REGION Network 5: Transfering
   RUNG wire#powerrail
      Contact( "R-201_Write_TO_T-102_DB".Transfering )
      Coil( "T-102_Read_FROM_R-201_DB".Transfering )
   END_RUNG
   // the same network as SCL:
   "T-102_Read_FROM_R-201_DB".Transfering := "R-201_Write_TO_T-102_DB".Transfering;
END_REGION

REGION Network 6: Filling Done
   RUNG wire#powerrail
      Contact( "R-201_Write_TO_T-102_DB".FillingDone )
      Coil( "T-102_Read_FROM_R-201_DB".FillingDone )
   END_RUNG
   // the same network as SCL:
   "T-102_Read_FROM_R-201_DB".FillingDone := "R-201_Write_TO_T-102_DB".FillingDone;
END_REGION

REGION Network 7: Aborting
   RUNG wire#powerrail
      Contact( "R-201_Write_TO_T-102_DB".Abort )
      Coil( "T-102_Read_FROM_R-201_DB".Aborting )
   END_RUNG
   // the same network as SCL:
   "T-102_Read_FROM_R-201_DB".Aborting := "R-201_Write_TO_T-102_DB".Abort;
END_REGION

REGION Network 8: Release Tank
   RUNG wire#powerrail
      Contact( "R-201_Write_TO_T-102_DB".ReleaseTank )
      Coil( "T-102_Read_FROM_R-201_DB".ReleaseTank )
   END_RUNG
   // the same network as SCL:
   "T-102_Read_FROM_R-201_DB".ReleaseTank := "R-201_Write_TO_T-102_DB".ReleaseTank;
END_REGION
END_FUNCTION

// folder: State MACHINE/1)Tanks/Tank T-102 (Y)/T-102 <---> R-202

FUNCTION "T-102_Signals_FROM_R-202" : Void   // FC70, LAD
{ S7_Optimized_Access := 'TRUE' }
VERSION : 0.1
BEGIN

REGION Network 1: Start Pouring Sequence
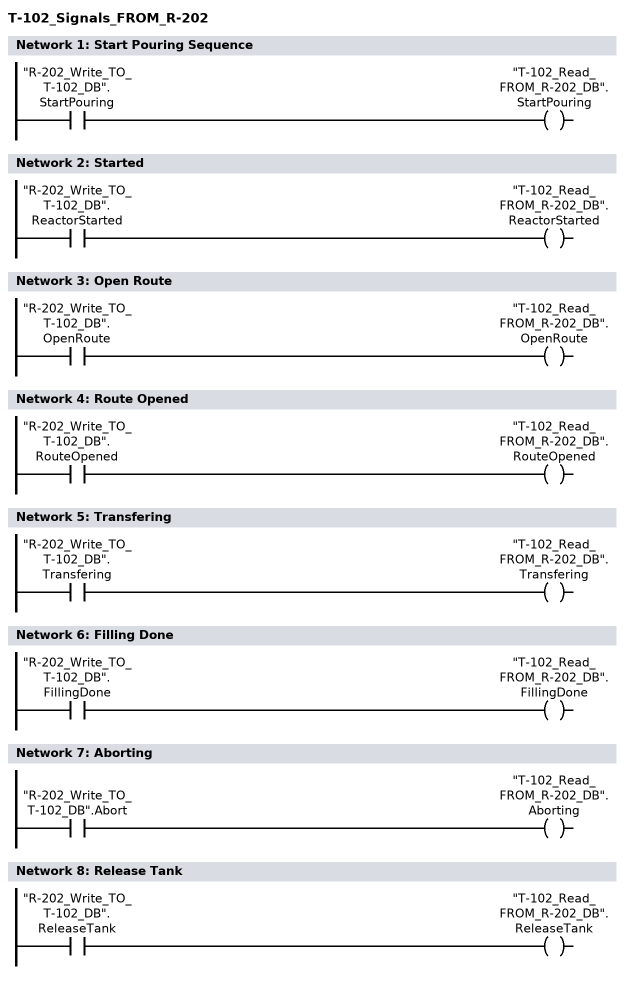
   RUNG wire#powerrail
      Contact( "R-202_Write_TO_T-102_DB".StartPouring )
      Coil( "T-102_Read_FROM_R-202_DB".StartPouring )
   END_RUNG
   // the same network as SCL:
   "T-102_Read_FROM_R-202_DB".StartPouring := "R-202_Write_TO_T-102_DB".StartPouring;
END_REGION

REGION Network 2: Started
   RUNG wire#powerrail
      Contact( "R-202_Write_TO_T-102_DB".ReactorStarted )
      Coil( "T-102_Read_FROM_R-202_DB".ReactorStarted )
   END_RUNG
   // the same network as SCL:
   "T-102_Read_FROM_R-202_DB".ReactorStarted := "R-202_Write_TO_T-102_DB".ReactorStarted;
END_REGION

REGION Network 3: Open Route
   RUNG wire#powerrail
      Contact( "R-202_Write_TO_T-102_DB".OpenRoute )
      Coil( "T-102_Read_FROM_R-202_DB".OpenRoute )
   END_RUNG
   // the same network as SCL:
   "T-102_Read_FROM_R-202_DB".OpenRoute := "R-202_Write_TO_T-102_DB".OpenRoute;
END_REGION

REGION Network 4: Route Opened
   RUNG wire#powerrail
      Contact( "R-202_Write_TO_T-102_DB".RouteOpened )
      Coil( "T-102_Read_FROM_R-202_DB".RouteOpened )
   END_RUNG
   // the same network as SCL:
   "T-102_Read_FROM_R-202_DB".RouteOpened := "R-202_Write_TO_T-102_DB".RouteOpened;
END_REGION

REGION Network 5: Transfering
   RUNG wire#powerrail
      Contact( "R-202_Write_TO_T-102_DB".Transfering )
      Coil( "T-102_Read_FROM_R-202_DB".Transfering )
   END_RUNG
   // the same network as SCL:
   "T-102_Read_FROM_R-202_DB".Transfering := "R-202_Write_TO_T-102_DB".Transfering;
END_REGION

REGION Network 6: Filling Done
   RUNG wire#powerrail
      Contact( "R-202_Write_TO_T-102_DB".FillingDone )
      Coil( "T-102_Read_FROM_R-202_DB".FillingDone )
   END_RUNG
   // the same network as SCL:
   "T-102_Read_FROM_R-202_DB".FillingDone := "R-202_Write_TO_T-102_DB".FillingDone;
END_REGION

REGION Network 7: Aborting
   RUNG wire#powerrail
      Contact( "R-202_Write_TO_T-102_DB".Abort )
      Coil( "T-102_Read_FROM_R-202_DB".Aborting )
   END_RUNG
   // the same network as SCL:
   "T-102_Read_FROM_R-202_DB".Aborting := "R-202_Write_TO_T-102_DB".Abort;
END_REGION

REGION Network 8: Release Tank
   RUNG wire#powerrail
      Contact( "R-202_Write_TO_T-102_DB".ReleaseTank )
      Coil( "T-102_Read_FROM_R-202_DB".ReleaseTank )
   END_RUNG
   // the same network as SCL:
   "T-102_Read_FROM_R-202_DB".ReleaseTank := "R-202_Write_TO_T-102_DB".ReleaseTank;
END_REGION
END_FUNCTION

// folder: State MACHINE/1)Tanks/Tank T-102 (Y)/T-102 <---> T-104

FUNCTION "T-102_Signals_FROM_T-104" : Void   // FC55, LAD
{ S7_Optimized_Access := 'TRUE' }
VERSION : 0.1
BEGIN

REGION Network 1: Start Sequence
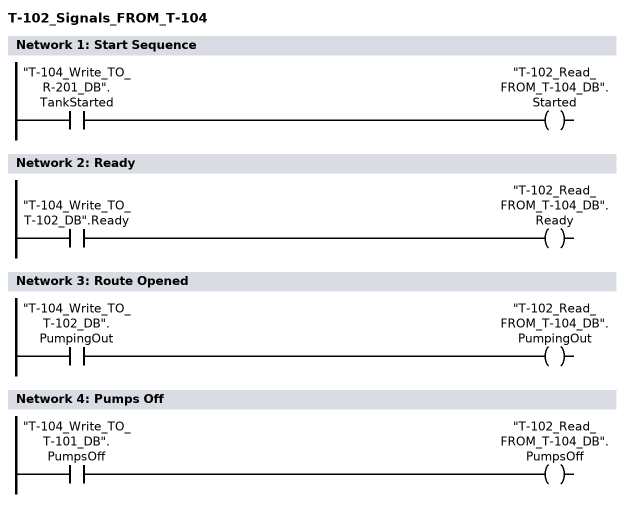
   RUNG wire#powerrail
      Contact( "T-104_Write_TO_R-201_DB".TankStarted )
      Coil( "T-102_Read_FROM_T-104_DB".Started )
   END_RUNG
   // the same network as SCL:
   "T-102_Read_FROM_T-104_DB".Started := "T-104_Write_TO_R-201_DB".TankStarted;
END_REGION

REGION Network 2: Ready
   RUNG wire#powerrail
      Contact( "T-104_Write_TO_T-102_DB".Ready )
      Coil( "T-102_Read_FROM_T-104_DB".Ready )
   END_RUNG
   // the same network as SCL:
   "T-102_Read_FROM_T-104_DB".Ready := "T-104_Write_TO_T-102_DB".Ready;
END_REGION

REGION Network 3: Route Opened
   RUNG wire#powerrail
      Contact( "T-104_Write_TO_T-102_DB".PumpingOut )
      Coil( "T-102_Read_FROM_T-104_DB".PumpingOut )
   END_RUNG
   // the same network as SCL:
   "T-102_Read_FROM_T-104_DB".PumpingOut := "T-104_Write_TO_T-102_DB".PumpingOut;
END_REGION

REGION Network 4: Pumps Off
   RUNG wire#powerrail
      Contact( "T-104_Write_TO_T-101_DB".PumpsOff )
      Coil( "T-102_Read_FROM_T-104_DB".PumpsOff )
   END_RUNG
   // the same network as SCL:
   "T-102_Read_FROM_T-104_DB".PumpsOff := "T-104_Write_TO_T-101_DB".PumpsOff;
END_REGION
END_FUNCTION

// folder: State MACHINE/1)Tanks/Tank T-103 (Cooling Tank)

FUNCTION_BLOCK "T-103_SEQ"   // FB33, GRAPH_PLUS
{ S7_Optimized_Access := 'TRUE' }
VERSION : 0.1
   VAR_INPUT
      OFF_SQ : Bool := false;   // Turn sequence off
      INIT_SQ : Bool := false;   // Set sequence to initial state
      ACK_EF : Bool := false;   // Acknowledge all errors and faults
   END_VAR
   VAR_OUTPUT
      S_NO : Int := 0;   // Step number
      S_MORE : Bool := false;   // More steps are available and can be shown in S_NO
      S_ACTIVE : Bool := false;   // Step indicated in S_NO is active
      ERR_FLT : Bool := false;   // Interlock or supervision group error
      AUTO_ON : Bool := false;   // Automatic mode is active
   END_VAR
   VAR
      STATE : Int;   // Current Step in Sequence
      Tank : Struct   // Reactor Ctrl
         IDLE : Bool;
         INITIALIZATION : Bool;   // Sequence initialization
         START : Bool;
         DONE_REACTING : Bool;
         COMPLETE : Bool;   // Reactor Complete Read only
         PARA : Bool;   // PARA load Batch side button
         ABORTING : Bool;   // Sequence about
         WAIT : Bool;   // Wating for Permissive read only
      END_STRUCT;
      TEMP : Struct
         TANKS_BATCH : Real;
         "EMPTY_LV_0%" : Real;
         "MIN_LV_20%" : Real;
         "MAX_LV_80%" : Real;
         "BELOW_32%" : Real;
         "Greater_8%" : Real;
         "PRE-ADD" : Real;
         X_SOL_SIZE : Real;
         Y_SOL_SIZE : Real;
         OFFSEt : Struct
            MAX : Real;
            MIN : Real;
         END_STRUCT;
      END_STRUCT;
      HMI_INFO : Array[0..12] of UInt;
      IF_PAR : G7_IfParPlus_V6;
      RT_DATA : G7_RTDataPlus_V6;   // Internal data area
      Abort : G7_TransitionPlus_V6;   // Transition structure
      Initialize : G7_TransitionPlus_V6;   // Transition structure
      Block : G7_TransitionPlus_V6;   // Transition structure
      Rdy : G7_TransitionPlus_V6;   // Transition structure
      Receive : G7_TransitionPlus_V6;   // Transition structure
      Centrifuge : G7_TransitionPlus_V6;   // Transition structure
      OpenR : G7_TransitionPlus_V6;   // Transition structure
      MinLevel : G7_TransitionPlus_V6;   // Transition structure
      DnTransf : G7_TransitionPlus_V6;   // Transition structure
      Cold : G7_TransitionPlus_V6;   // Transition structure
      POff : G7_TransitionPlus_V6;   // Transition structure
      ClsR : G7_TransitionPlus_V6;   // Transition structure
      DnClng : G7_TransitionPlus_V6;   // Transition structure
      TrSt : G7_TransitionPlus_V6;   // Transition structure
      ROpn : G7_TransitionPlus_V6;   // Transition structure
      Tng : G7_TransitionPlus_V6;   // Transition structure
      ClsFR : G7_TransitionPlus_V6;   // Transition structure
      DnT : G7_TransitionPlus_V6;   // Transition structure
      Init : G7_TransitionPlus_V6;   // Transition structure
      SAut : G7_TransitionPlus_V6;   // Transition structure
      SIn : G7_TransitionPlus_V6;   // Transition structure
      Initd : G7_TransitionPlus_V6;   // Transition structure
      BskFull : G7_TransitionPlus_V6;   // Transition structure
      FeelerRet : G7_TransitionPlus_V6;   // Transition structure
      Ab : G7_TransitionPlus_V6;   // Transition structure
      AbortOn : G7_TransitionPlus_V6;   // Transition structure
      DneAbort : G7_TransitionPlus_V6;   // Transition structure
      Idle : G7_StepPlus_V6;   // Step structure
      Ready : G7_StepPlus_V6;   // Step structure
      SelectSeq : G7_StepPlus_V6;   // Step structure
      Started : G7_StepPlus_V6;   // Step structure
      Filling : G7_StepPlus_V6;   // Step structure
      "Filling/Tansfer" : G7_StepPlus_V6;   // Step structure
      Wait_Temp : G7_StepPlus_V6;   // Step structure
      PmpOff : G7_StepPlus_V6;   // Step structure
      CloseRecirc : G7_StepPlus_V6;   // Step structure
      "USER Ready" : G7_StepPlus_V6;   // Step structure
      ReadyToTransf : G7_StepPlus_V6;   // Step structure
      RouteOpened : G7_StepPlus_V6;   // Step structure
      Transfering : G7_StepPlus_V6;   // Step structure
      CloseFeedRoute : G7_StepPlus_V6;   // Step structure
      DoneTrnf : G7_StepPlus_V6;   // Step structure
      Idle_Init : G7_StepPlus_V6;   // Step structure
      SetAuto : G7_StepPlus_V6;   // Step structure
      SetInitial : G7_StepPlus_V6;   // Step structure
      Done_Init : G7_StepPlus_V6;   // Step structure
      AbortStarting : G7_StepPlus_V6;   // Step structure
      Aborting : G7_StepPlus_V6;   // Step structure
      Abort_Done : G7_StepPlus_V6;   // Step structure
      SINI : Array[0..5] of USInt;
      LSTT : Array[0..26] of USInt;
      ATAJ : Array[0..26] of USInt;
      ATAB : Array[0..26] of USInt;
      PSTT : Array[0..26] of USInt;
      NSTT : Array[0..26] of USInt;
      ASSJ : Array[0..21] of USInt;
      ASSB : Array[0..21] of USInt;
      PTTS : Array[0..21] of USInt;
      NTTS : Array[0..21] of USInt;
      SW_SQTS : Array[0..21] of USInt;
      SWITCH : Array[0..6] of USInt;
      TVX : Array[0..13] of USInt;
      TTX : Array[0..13] of USInt;
      TSX : Array[0..5] of USInt;
      S00X : Array[0..5] of USInt;
      SOFFX : Array[0..5] of USInt;
      SONX : Array[0..5] of USInt;
      SAX : Array[0..5] of USInt;
      SERRX : Array[0..22] of USInt;
      SMX : Array[0..22] of USInt;
      S0X : Array[0..22] of USInt;
      S1X : Array[0..22] of USInt;
      IL_ALARM_INST : Diag_Alarm;
      SUP_ALARM_INST : Diag_Alarm;
      STEP_TIME_ALARM_INST : Diag_Alarm;
      IEC_TIMER_INST : IEC_TIMER;
      TRANSACTION_FLAG : Bool := false;
   END_VAR
   VAR CONSTANT
      "Single R-201 T-101 seq done" : Int := 214;
      "Single R-201 T-102 seq done" : Int := 218;
   END_VAR
   // SINI[0] := 2;
   // LSTT[0] := 19;
   // NSTT[0] := 19;
   // PTTS[0] := 255;
   // TVX[0] := 16#1;
   // TTX[0] := 16#1;
   // TSX[0] := 16#1;
   // S00X[0] := 16#1;
   // SOFFX[0] := 16#1;
   // SONX[0] := 16#1;
   // SAX[0] := 16#1;
   // SERRX[0] := 16#1;
   // SMX[0] := 16#1;
   // S0X[0] := 16#1;
   // S1X[0] := 16#1;
   // LSTT[1] := 15;
   // LSTT[2] := 255;
   // LSTT[3] := 255;
   // LSTT[4] := 3;
   // LSTT[5] := 10;
   // LSTT[6] := 255;
   // LSTT[7] := 255;
   // LSTT[8] := 255;
   // LSTT[9] := 255;
   // LSTT[10] := 255;
   // LSTT[11] := 255;
   // LSTT[21] := 1;
   // LSTT[13] := 255;
   // LSTT[14] := 255;
   // LSTT[15] := 255;
   // LSTT[16] := 255;
   // LSTT[20] := 255;
   // LSTT[23] := 10;
   // LSTT[19] := 255;
   // LSTT[22] := 10;
   // ATAJ[1] := 1;
   // ATAJ[2] := 2;
   // ATAJ[3] := 3;
   // ATAJ[4] := 4;
   // ATAJ[5] := 5;
   // ATAJ[6] := 6;
   // ATAJ[7] := 7;
   // ATAJ[8] := 8;
   // ATAJ[9] := 9;
   // ATAJ[10] := 10;
   // ATAJ[11] := 11;
   // ATAJ[12] := 12;
   // ATAJ[13] := 13;
   // ATAJ[14] := 14;
   // ATAJ[15] := 15;
   // ATAJ[16] := 16;
   // ATAJ[17] := 17;
   // ATAJ[18] := 18;
   // ATAJ[19] := 19;
   // ATAJ[20] := 20;
   // ATAJ[21] := 21;
   // ATAJ[22] := 22;
   // ATAJ[23] := 23;
   // ATAJ[24] := 24;
   // ATAB[1] := 2;
   // ATAB[10] := 10;
   // ATAB[3] := 3;
   // ATAB[4] := 5;
   // ATAB[5] := 4;
   // ATAB[6] := 6;
   // ATAB[7] := 7;
   // ATAB[8] := 8;
   // ATAB[12] := 12;
   // ATAB[11] := 11;
   // ATAB[13] := 13;
   // ATAB[14] := 14;
   // ATAB[15] := 22;
   // ATAB[16] := 16;
   // ATAB[17] := 17;
   // ATAB[18] := 18;
   // ATAB[21] := 21;
   // ATAB[22] := 23;
   // ATAB[23] := 15;
   // ATAB[24] := 24;
   // ATAB[0] := 1;
   // PSTT[10] := 7;
   // PSTT[16] := 13;
   // PSTT[3] := 1;
   // PSTT[4] := 2;
   // PSTT[5] := 2;
   // PSTT[6] := 3;
   // PSTT[7] := 4;
   // PSTT[12] := 9;
   // PSTT[11] := 8;
   // PSTT[13] := 10;
   // PSTT[14] := 11;
   // PSTT[17] := 14;
   // PSTT[18] := 15;
   // PSTT[19] := 16;
   // PSTT[20] := 17;
   // PSTT[21] := 18;
   // PSTT[22] := 12;
   // PSTT[23] := 12;
   // PSTT[24] := 19;
   // NSTT[1] := 15;
   // NSTT[2] := 1;
   // NSTT[3] := 2;
   // NSTT[4] := 3;
   // NSTT[5] := 10;
   // NSTT[6] := 4;
   // NSTT[7] := 5;
   // NSTT[8] := 6;
   // NSTT[9] := 7;
   // NSTT[10] := 8;
   // NSTT[11] := 9;
   // NSTT[21] := 1;
   // NSTT[13] := 11;
   // NSTT[14] := 12;
   // NSTT[15] := 13;
   // NSTT[16] := 14;
   // NSTT[20] := 18;
   // NSTT[23] := 10;
   // NSTT[19] := 17;
   // NSTT[22] := 10;
   // ASSJ[1] := 1;
   // ASSJ[2] := 2;
   // ASSJ[3] := 3;
   // ASSJ[4] := 4;
   // ASSJ[5] := 5;
   // ASSJ[6] := 6;
   // ASSJ[7] := 7;
   // ASSJ[8] := 8;
   // ASSJ[9] := 9;
   // ASSJ[10] := 10;
   // ASSJ[11] := 11;
   // ASSJ[12] := 12;
   // ASSJ[13] := 13;
   // ASSJ[14] := 14;
   // ASSJ[15] := 15;
   // ASSJ[16] := 16;
   // ASSJ[17] := 17;
   // ASSJ[18] := 18;
   // ASSJ[19] := 19;
   // ASSJ[20] := 20;
   // ASSJ[21] := 21;
   // ASSB[1] := 1;
   // ASSB[2] := 2;
   // ASSB[3] := 3;
   // ASSB[4] := 4;
   // ASSB[5] := 5;
   // ASSB[6] := 6;
   // ASSB[7] := 7;
   // ASSB[8] := 8;
   // ASSB[9] := 9;
   // ASSB[10] := 10;
   // ASSB[11] := 11;
   // ASSB[12] := 12;
   // ASSB[13] := 13;
   // ASSB[14] := 14;
   // ASSB[15] := 15;
   // ASSB[16] := 16;
   // ASSB[17] := 17;
   // ASSB[18] := 18;
   // ASSB[19] := 19;
   // ASSB[20] := 20;
   // ASSB[21] := 21;
   // PTTS[4] := 6;
   // PTTS[3] := 255;
   // PTTS[5] := 7;
   // PTTS[6] := 8;
   // PTTS[7] := 9;
   // PTTS[8] := 10;
   // PTTS[9] := 11;
   // PTTS[10] := 255;
   // PTTS[11] := 13;
   // PTTS[12] := 14;
   // PTTS[13] := 15;
   // PTTS[14] := 16;
   // PTTS[15] := 255;
   // PTTS[16] := 18;
   // PTTS[17] := 19;
   // PTTS[18] := 20;
   // PTTS[19] := 255;
   // PTTS[20] := 24;
   // PTTS[21] := 25;
   // SW_SQTS[4] := 2;
   // NTTS[2] := 4;
   // NTTS[3] := 6;
   // NTTS[4] := 7;
   // NTTS[5] := 8;
   // NTTS[6] := 9;
   // NTTS[7] := 10;
   // NTTS[8] := 11;
   // NTTS[9] := 12;
   // NTTS[10] := 13;
   // NTTS[11] := 14;
   // NTTS[12] := 15;
   // NTTS[13] := 16;
   // NTTS[14] := 17;
   // NTTS[15] := 18;
   // NTTS[16] := 19;
   // NTTS[17] := 20;
   // NTTS[18] := 21;
   // NTTS[19] := 24;
   // NTTS[20] := 25;
   // NTTS[21] := 26;
   // SW_SQTS[5] := 2;
   // SW_SQTS[8] := 2;
   // SW_SQTS[9] := 2;
   // SW_SQTS[10] := 3;
   // SW_SQTS[11] := 3;
   // SW_SQTS[12] := 3;
   // SW_SQTS[13] := 4;
   // SW_SQTS[14] := 4;
   // SW_SQTS[15] := 5;
   // SW_SQTS[16] := 5;
   // SW_SQTS[17] := 5;
   // SW_SQTS[18] := 5;
   // SW_SQTS[19] := 6;
   // SW_SQTS[20] := 6;
   // SW_SQTS[21] := 6;
   // SWITCH[3] := 124;
   // SWITCH[0] := 124;
   // SWITCH[2] := 254;
   // SWITCH[4] := 254;
   // PTTS[2] := 3;
   // SW_SQTS[3] := 2;
   // SWITCH[1] := 254;
   // SW_SQTS[2] := 1;
   // ATAB[20] := 20;
   // PSTT[9] := 6;
   // PTTS[1] := 2;
   // NTTS[1] := 3;
   // SW_SQTS[1] := 1;
   // SINI[3] := 255;
   // ATAB[19] := 19;
   // PSTT[15] := 12;
   // SW_SQTS[7] := 2;
   // SW_SQTS[6] := 2;
   // SINI[2] := 255;
   // SINI[4] := 255;
   // SINI[5] := 255;
   // LSTT[18] := 255;
   // ATAB[9] := 9;
   // PSTT[8] := 5;
   // NSTT[18] := 16;
   // LSTT[12] := 10;
   // NSTT[12] := 10;
   // LSTT[24] := 255;
   // LSTT[25] := 255;
   // ATAJ[25] := 25;
   // ATAJ[26] := 26;
   // ATAB[25] := 25;
   // ATAB[26] := 26;
   // PSTT[25] := 20;
   // PSTT[26] := 21;
   // NSTT[24] := 20;
   // NSTT[25] := 21;
   // SWITCH[5] := 254;
BEGIN
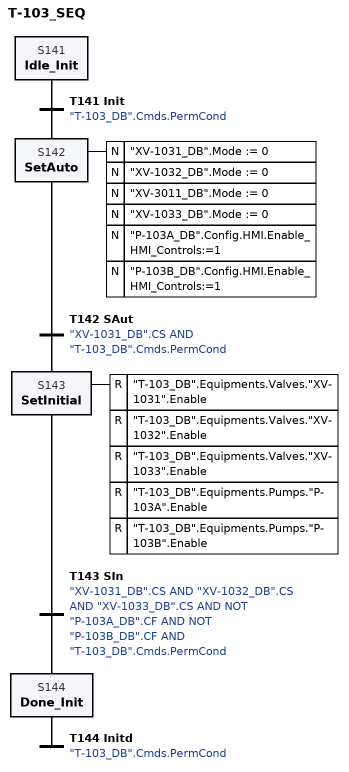
   // permanent pre-instructions
   NETWORK 1
      "T-103_Signals_FROM_R-201"();
      "T-103_Signals_FROM_R-202"();
      "T-103_Signals_FROM_Centrifuge"();
      "T-103_SignalsInExchange"();
      "T-103_SEQ_FC"();

   // sequencer 1
   STEP SetInitial:   // S143, max time T#10S, warning time T#7S
      // Initialize Batch sequence
              R    "T-103_DB".Equipments.Valves."XV-1031".Enable
              R    "T-103_DB".Equipments.Valves."XV-1032".Enable
              R    "T-103_DB".Equipments.Valves."XV-1033".Enable
              R    "T-103_DB".Equipments.Pumps."P-103A".Enable
              R    "T-103_DB".Equipments.Pumps."P-103B".Enable
   END_STEP
   TRANSITION SIn FROM SetInitial TO Done_Init   // T143: OFF: P-101A/B
      := "XV-1031_DB".CS AND "XV-1032_DB".CS AND "XV-1033_DB".CS AND NOT "P-103A_DB".CF AND NOT "P-103B_DB".CF AND "T-103_DB".Cmds.PermCond;
   END_TRANSITION
   STEP Idle_Init:   // S141, max time T#10S, warning time T#7S
   END_STEP
   TRANSITION Init FROM Idle_Init TO SetAuto   // T141
      := "T-103_DB".Cmds.PermCond;
   END_TRANSITION
   STEP SetAuto:   // S142, max time T#10S, warning time T#7S
      // Initialize Batch sequence
              N    "XV-1031_DB".Mode := 0
              N    "XV-1032_DB".Mode := 0
              N    "XV-3011_DB".Mode := 0
              N    "XV-1033_DB".Mode := 0
              N    "P-103A_DB".Config.HMI.Enable_HMI_Controls:=1
              N    "P-103B_DB".Config.HMI.Enable_HMI_Controls:=1
   END_STEP
   TRANSITION SAut FROM SetAuto TO SetInitial   // T142: CLOSED: XV-1041 XV-1011 XV-1013OFF: VFD-1011 P-101A P-101BZERO: FT-1041 Totalizer
      := "XV-1031_DB".CS AND "T-103_DB".Cmds.PermCond;
   END_TRANSITION
   STEP Done_Init:   // S144, max time T#10S, warning time T#7S
   END_STEP
   TRANSITION Initd FROM Done_Init TO ?   // T144
      := "T-103_DB".Cmds.PermCond;
   END_TRANSITION

   // permanent post-instructions
   NETWORK 1
      "T-103_SignalsOutExchange"();
      "T-103_FC_Outputs"();
END_FUNCTION_BLOCK

FUNCTION "T-103_SignalsInExchange" : Void   // FC41, LAD
{ S7_Optimized_Access := 'TRUE' }
VERSION : 0.1
BEGIN

REGION Network 1: Start Receiving (Receive)
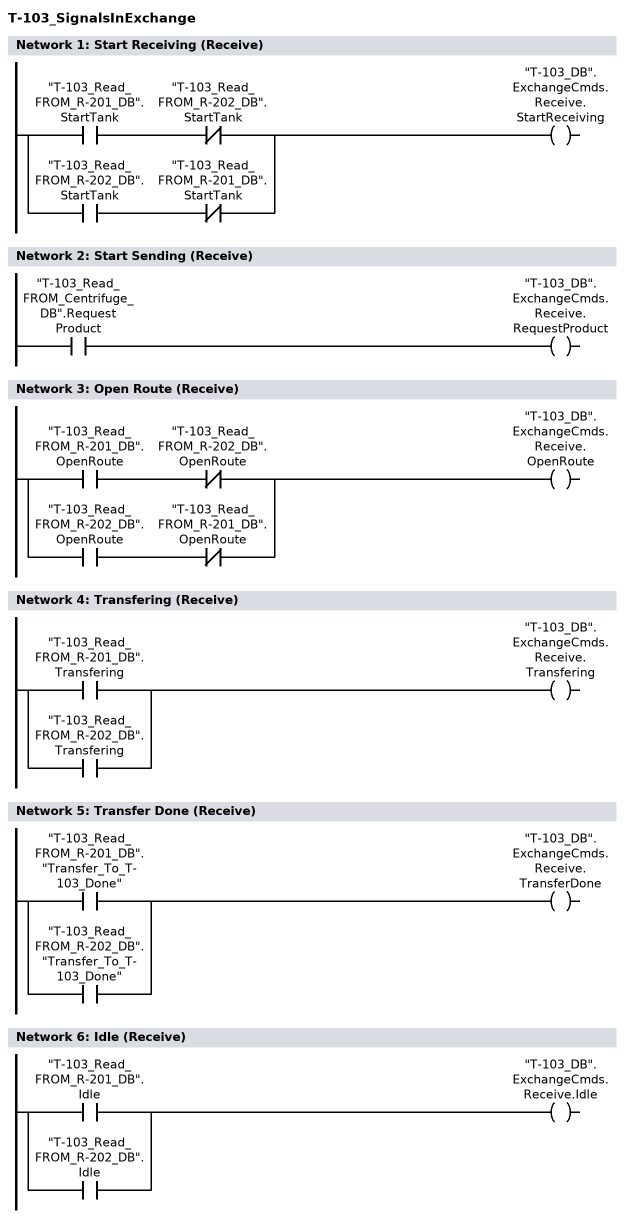
   RUNG wire#powerrail
      Contact( "T-103_Read_FROM_R-201_DB".StartTank )
      I_Contact( "T-103_Read_FROM_R-202_DB".StartTank )
      wire#w1
      Coil( "T-103_DB".ExchangeCmds.Receive.StartReceiving )
   END_RUNG
   RUNG wire#powerrail
      Contact( "T-103_Read_FROM_R-202_DB".StartTank )
      I_Contact( "T-103_Read_FROM_R-201_DB".StartTank )
   END_RUNG wire#w1
   // the same network as SCL:
   "T-103_DB".ExchangeCmds.Receive.StartReceiving := ("T-103_Read_FROM_R-201_DB".StartTank AND NOT "T-103_Read_FROM_R-202_DB".StartTank) OR ("T-103_Read_FROM_R-202_DB".StartTank AND NOT "T-103_Read_FROM_R-201_DB".StartTank);
END_REGION

REGION Network 2: Start Sending (Receive)
   RUNG wire#powerrail
      Contact( "T-103_Read_FROM_Centrifuge_DB".RequestProduct )
      Coil( "T-103_DB".ExchangeCmds.Receive.RequestProduct )
   END_RUNG
   // the same network as SCL:
   "T-103_DB".ExchangeCmds.Receive.RequestProduct := "T-103_Read_FROM_Centrifuge_DB".RequestProduct;
END_REGION

REGION Network 3: Open Route (Receive)
   RUNG wire#powerrail
      Contact( "T-103_Read_FROM_R-201_DB".OpenRoute )
      I_Contact( "T-103_Read_FROM_R-202_DB".OpenRoute )
      wire#w1
      Coil( "T-103_DB".ExchangeCmds.Receive.OpenRoute )
   END_RUNG
   RUNG wire#powerrail
      Contact( "T-103_Read_FROM_R-202_DB".OpenRoute )
      I_Contact( "T-103_Read_FROM_R-201_DB".OpenRoute )
   END_RUNG wire#w1
   // the same network as SCL:
   "T-103_DB".ExchangeCmds.Receive.OpenRoute := ("T-103_Read_FROM_R-201_DB".OpenRoute AND NOT "T-103_Read_FROM_R-202_DB".OpenRoute) OR ("T-103_Read_FROM_R-202_DB".OpenRoute AND NOT "T-103_Read_FROM_R-201_DB".OpenRoute);
END_REGION

REGION Network 4: Transfering (Receive)
   RUNG wire#powerrail
      Contact( "T-103_Read_FROM_R-201_DB".Transfering )
      wire#w1
      Coil( "T-103_DB".ExchangeCmds.Receive.Transfering )
   END_RUNG
   RUNG wire#powerrail
      Contact( "T-103_Read_FROM_R-202_DB".Transfering )
   END_RUNG wire#w1
   // the same network as SCL:
   "T-103_DB".ExchangeCmds.Receive.Transfering := "T-103_Read_FROM_R-201_DB".Transfering OR "T-103_Read_FROM_R-202_DB".Transfering;
END_REGION

REGION Network 5: Transfer Done (Receive)
   RUNG wire#powerrail
      Contact( "T-103_Read_FROM_R-201_DB"."Transfer_To_T-103_Done" )
      wire#w1
      Coil( "T-103_DB".ExchangeCmds.Receive.TransferDone )
   END_RUNG
   RUNG wire#powerrail
      Contact( "T-103_Read_FROM_R-202_DB"."Transfer_To_T-103_Done" )
   END_RUNG wire#w1
   // the same network as SCL:
   "T-103_DB".ExchangeCmds.Receive.TransferDone := "T-103_Read_FROM_R-201_DB"."Transfer_To_T-103_Done" OR "T-103_Read_FROM_R-202_DB"."Transfer_To_T-103_Done";
END_REGION

REGION Network 6: Idle (Receive)
   RUNG wire#powerrail
      Contact( "T-103_Read_FROM_R-201_DB".Idle )
      wire#w1
      Coil( "T-103_DB".ExchangeCmds.Receive.Idle )
   END_RUNG
   RUNG wire#powerrail
      Contact( "T-103_Read_FROM_R-202_DB".Idle )
   END_RUNG wire#w1
   // the same network as SCL:
   "T-103_DB".ExchangeCmds.Receive.Idle := "T-103_Read_FROM_R-201_DB".Idle OR "T-103_Read_FROM_R-202_DB".Idle;
END_REGION
END_FUNCTION

FUNCTION "T-103_FC_Outputs" : Void   // FC82, SCL
{ S7_Optimized_Access := 'TRUE' }
VERSION : 0.1
   VAR_TEMP
      Pump_A : Struct
         Cond_01 : Bool;   // Condition 01
         Cond_02 : Bool;
         Cond_03 : Bool;   // Condition 03
      END_STRUCT;
      Pump_B : Struct
         Cond_01 : Bool;   // Condition 01
         Cond_02 : Bool;   // Condition 02
         Cond_03 : Bool;   // Condition 03
      END_STRUCT;
      Motor : Struct
         Cond_01 : Bool;   // Condition 01
         Cond_02 : Bool;   // Condition 02
         Cond_03 : Bool;   // Condition 03
      END_STRUCT;
      XV : Struct
         "1032" : Bool;
         "1031" : Bool;
         "3011" : Bool;
         "1033" : Bool;
      END_STRUCT;
   END_VAR
BEGIN
   //****** Equipmens Activation*******
   //
   //**************************************************************
   //IF "AlwaysFALSE" THEN

       //***********************************************Tank Outlet Valve**********************************************************************
       IF "XV-1032_DB".Mode = 0 THEN
           "T-103_DB".Equipments.Valves."XV-1032".CmdOn := "T-103_DB".Equipments.Valves."XV-1032".Enable AND NOT "T-103_DB".Cmds.Hold;
           //Delay Off To avoid Overpressure the Lines
           #XV."1032" := "T-103_DB".Equipments.Valves."XV-1032".CmdOn;
           "T-103_Aux_DB".Timer."XV-1032".TOF(IN := #XV."1032",
                                              PT := "T-103_Aux_DB".Constants.CmdDelay);
           //Command to the Valve
           IF "T-103_Aux_DB".Timer."XV-1032".Q THEN
               "XV-1032_DB".CMD := 2;
           ELSE
               "XV-1032_DB".CMD := 1;
           END_IF;
           "T-103_DB".Equipments.Valves."XV-1032".TurningOff := NOT "T-103_DB".Equipments.Valves."XV-1032".CmdOn AND "T-103_Aux_DB".Timer."XV-1032".Q;
       END_IF;
       //***********************************************Tank Inlet Valve**********************************************************************
       IF "XV-1031_DB".Mode = 0 THEN
           "T-103_DB".Equipments.Valves."XV-1031".CmdOn := "T-103_DB".Equipments.Valves."XV-1031".Enable AND NOT "T-103_DB".Cmds.Hold;
           //Delay Off To avoid Overpressure the Lines
           #XV."1031" := "T-103_DB".Equipments.Valves."XV-1031".CmdOn;
           "T-103_Aux_DB".Timer."XV-1031".TOF(IN := #XV."1031",
                                              PT := "T-103_Aux_DB".Constants.CmdDelay);
           IF "T-103_Aux_DB".Timer."XV-1031".Q THEN
               "XV-1031_DB".CMD := 2;
           ELSE
               "XV-1031_DB".CMD := 1;
           END_IF;
           "T-103_DB".Equipments.Valves."XV-1031".TurningOff := NOT "T-103_DB".Equipments.Valves."XV-1031".CmdOn AND "T-103_Aux_DB".Timer."XV-1031".Q;
       END_IF;
       ////***********************************************Recirculate valve**********************************************************************
       IF "XV-1033_DB".Mode = 0 THEN
           "T-103_DB".Equipments.Valves."XV-1033".CmdOn := "T-103_DB".Equipments.Valves."XV-1033".Enable AND NOT "T-103_DB".Cmds.Hold;
           //Delay Off To avoid Overpressure the Lines
           #XV."1033" := "T-103_DB".Equipments.Valves."XV-1033".CmdOn;
           "T-103_Aux_DB".Timer."XV-1033".TOF(IN := #XV."1033",
                                              PT := "T-103_Aux_DB".Constants.CmdDelay);
           IF "T-103_Aux_DB".Timer."XV-1033".Q THEN
               "XV-1033_DB".CMD := 2;
           ELSE
               "XV-1033_DB".CMD := 1;
           END_IF;
           "T-103_DB".Equipments.Valves."XV-1033".TurningOff := NOT "T-103_DB".Equipments.Valves."XV-1033".CmdOn AND "T-103_Aux_DB".Timer."XV-1033".Q;
       END_IF;
       //***********************************************T-103 Pump A**********************************************************************
       // Condition to CmdOn "On Command" 
       IF "P-103A_DB".Config.HMI.Enable_HMI_Controls = 1 THEN
           #Pump_A.Cond_01 := "T-103_DB".Equipments.Pumps."P-103A".Enable AND ("T-103_DB".PmpSel."P-103AB" = 1 OR "T-103_DB".PmpSel."P-103AB" = 3);
           #Pump_A.Cond_02 := "T-103_Read_FROM_Centrifuge_DB".RouteOpened AND "T-103_Write_TO_Centrifuge_DB".RouteOpened; //Route Open to sent to Centrifuge
           #Pump_A.Cond_03 := "XV-1033_DB".OS AND "XV-1032_DB".OS AND "XV-3011_DB".CS; //Route open to Recirculate
           "T-103_DB".Equipments.Pumps."P-103A".CmdOn := #Pump_A.Cond_01 AND (#Pump_A.Cond_02 OR #Pump_A.Cond_03);
           //**********Commands to the Pumps
           IF "T-103_DB".Equipments.Pumps."P-103A".CmdOn THEN
               "P-103A_DB".Stop_CMD := False;
               "P-103A_DB".Start_CMD := true;
               "P-103A_DB".ON := TRUE;
               "P-103A_DB".OFF := FALSE;
           ELSE
               "P-103A_DB".Stop_CMD := TRUE;
               "P-103A_DB".Start_CMD := FALSE;
               "P-103A_DB".ON := FALSE;
               "P-103A_DB".OFF := TRUE;
           END_IF;

           //*****Pressure Protection******

       END_IF;
       //***********************************************T-103 Pump B**********************************************************************
       // Condition to CmdOn "On Command" 
       IF "P-103B_DB".Config.HMI.Enable_HMI_Controls = 1 THEN
           #Pump_B.Cond_01 := "T-103_DB".Equipments.Pumps."P-103B".Enable AND ("T-103_DB".PmpSel."P-103AB" = 2 OR "T-103_DB".PmpSel."P-103AB" = 3);
           #Pump_B.Cond_02 := "T-103_Read_FROM_Centrifuge_DB".RouteOpened AND "T-103_Write_TO_Centrifuge_DB".RouteOpened; //Route Open to sent to Centrifuge
           #Pump_B.Cond_03 := "XV-1033_DB".OS AND "XV-1032_DB".OS AND "XV-3011_DB".CS; //Route open to Recirculate
           "T-103_DB".Equipments.Pumps."P-103B".CmdOn := #Pump_B.Cond_01 AND (#Pump_B.Cond_02 OR #Pump_B.Cond_03);
           //**********Commands to the Pumps
           IF "T-103_DB".Equipments.Pumps."P-103B".CmdOn THEN
               "P-103B_DB".Stop_CMD := False;
               "P-103B_DB".Start_CMD := true;
               "P-103B_DB".ON := TRUE;
               "P-103B_DB".OFF := FALSE;
           ELSE
               "P-103B_DB".Stop_CMD := TRUE;
               "P-103B_DB".Start_CMD := FALSE;
               "P-103B_DB".ON := FALSE;
               "P-103B_DB".OFF := TRUE;
           END_IF;
       END_IF;

       //***********************************************Mixer********************************************************************
       IF "VFD-T103_DB".HMI.Controls.Mode = 2 THEN
           #Motor.Cond_01 := "T-103_DB".Equipments.VFD."VFD-T103".Enable;
           "T-103_DB".Equipments.VFD."VFD-T103".CmdOn := #Motor.Cond_01 AND NOT "T-103_DB".Cmds.Hold AND NOT "T-103_DB".Status.Aborting;
           IF "T-103_DB".Equipments.VFD."VFD-T103".CmdOn THEN
               "VFD-T103_DB".PLCCommand := TRUE;
           ELSE
               "VFD-T103_DB".PLCCommand := FALSE;
           END_IF;
       END_IF;
       //END_IF;


   //END_IF;


   //****interlocks to reactor*****// Modification mode to transfer from Reactor to Centrifuge passing for T-103
       "T-103_DB".ExchangeCmds.Send.RouteOpened := "XV-1031_DB".OS AND "T-103_Read_FROM_Centrifuge_DB".RouteOpened; //Receive Material from Reactor.
   //*****Interlocks to Centrifuge*****//
   "T-103_Write_TO_Centrifuge_DB".RouteOpened := "XV-1032_DB".OS AND "XV-1033_DB".CS; //Send Material to Centrifuge
   "T-103_Write_TO_Centrifuge_DB".Transfering := ("XV-1032_DB".OS  AND "XV-1033_DB".CS) AND (("P-103A_DB".CF AND ("PT-103A_DB".SAI > 0.2)) OR ("P-103B_DB".CF AND ("PT-103B_DB".SAI > 0.2)));
   "T-103_Write_TO_Centrifuge_DB".Pumps_OFF := NOT "P-103A_DB".CF AND NOT "P-103B_DB".CF;

   //***************Valves Status***************//
   "T-103_Aux_DB"."Bool".TOff := "T-103_DB".Equipments.Valves."XV-1032".TurningOff OR "T-103_DB".Equipments.Valves."XV-1031".TurningOff OR "T-103_DB".Equipments.Valves."XV-3011".TurningOff OR "T-103_DB".Equipments.Valves."XV-1033".TurningOff;
   //*********************************Timers***********************************************************
   //Delay to Start Recirculation when transfering from Reactors.
   "T-103_Aux_DB"."Bool".StartRecirD_Enab := "T-103_DB".Status.Step = 22 AND "T-103_DB".ExchangeCmds.Receive.Transfering;
END_FUNCTION

FUNCTION "T-103_SignalsOutExchange" : Void   // FC89, LAD
{ S7_Optimized_Access := 'TRUE' }
VERSION : 0.1
BEGIN

REGION Network 1: Started (Send)
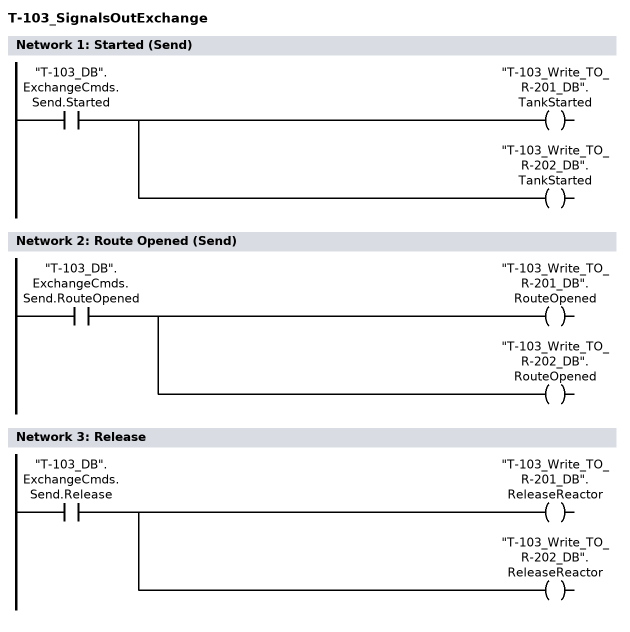
   RUNG wire#powerrail
      Contact( "T-103_DB".ExchangeCmds.Send.Started )
      wire#w1
      Coil( "T-103_Write_TO_R-201_DB".TankStarted )
   END_RUNG
   RUNG wire#w1
      Coil( "T-103_Write_TO_R-202_DB".TankStarted )
   END_RUNG
   // the same network as SCL:
   "T-103_Write_TO_R-201_DB".TankStarted := "T-103_DB".ExchangeCmds.Send.Started;
   "T-103_Write_TO_R-202_DB".TankStarted := "T-103_DB".ExchangeCmds.Send.Started;
END_REGION

REGION Network 2: Route Opened (Send)
   RUNG wire#powerrail
      Contact( "T-103_DB".ExchangeCmds.Send.RouteOpened )
      wire#w1
      Coil( "T-103_Write_TO_R-201_DB".RouteOpened )
   END_RUNG
   RUNG wire#w1
      Coil( "T-103_Write_TO_R-202_DB".RouteOpened )
   END_RUNG
   // the same network as SCL:
   "T-103_Write_TO_R-201_DB".RouteOpened := "T-103_DB".ExchangeCmds.Send.RouteOpened;
   "T-103_Write_TO_R-202_DB".RouteOpened := "T-103_DB".ExchangeCmds.Send.RouteOpened;
END_REGION

REGION Network 3: Release
   RUNG wire#powerrail
      Contact( "T-103_DB".ExchangeCmds.Send.Release )
      wire#w1
      Coil( "T-103_Write_TO_R-201_DB".ReleaseReactor )
   END_RUNG
   RUNG wire#w1
      Coil( "T-103_Write_TO_R-202_DB".ReleaseReactor )
   END_RUNG
   // the same network as SCL:
   "T-103_Write_TO_R-201_DB".ReleaseReactor := "T-103_DB".ExchangeCmds.Send.Release;
   "T-103_Write_TO_R-202_DB".ReleaseReactor := "T-103_DB".ExchangeCmds.Send.Release;
END_REGION
END_FUNCTION

FUNCTION "T-103_SEQ_FC" : Void   // FC90, LAD
{ S7_Optimized_Access := 'TRUE' }
VERSION : 0.1
   VAR_TEMP   // added for the SCL form of the ladder/FBD networks
      _w1 : Bool;
      _w2 : Bool;
      _w3 : Bool;
   END_VAR
BEGIN

REGION Network 2: Abort
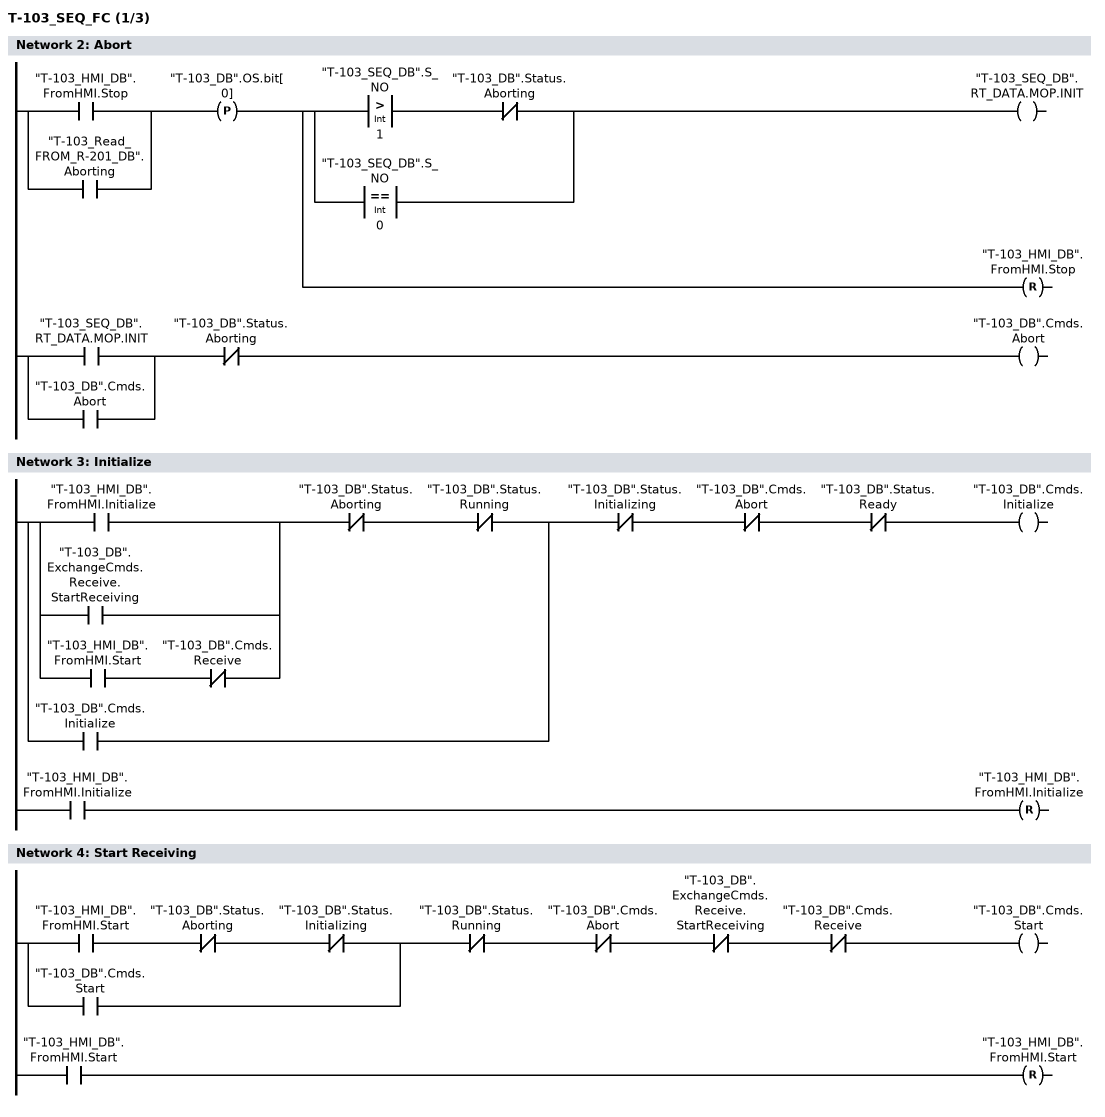
   RUNG wire#powerrail
      Contact( "T-103_HMI_DB".FromHMI.Stop )
      wire#w1
      P_Trig( "T-103_DB".OS.bit[0] )
      wire#w2
      { S7_Templates := "SrcType := Int" } GT_Contact(in1 := "T-103_SEQ_DB".S_NO, in2 := 1)
      I_Contact( "T-103_DB".Status.Aborting )
      wire#w3
      Coil( "T-103_SEQ_DB".RT_DATA.MOP.INIT )
   END_RUNG
   RUNG wire#powerrail
      Contact( "T-103_Read_FROM_R-201_DB".Aborting )
   END_RUNG wire#w1
   RUNG wire#w2
      { S7_Templates := "SrcType := Int" } EQ_Contact(in1 := "T-103_SEQ_DB".S_NO, in2 := 0)
   END_RUNG wire#w3
   RUNG wire#w2
      R_Coil( "T-103_HMI_DB".FromHMI.Stop )
   END_RUNG
   RUNG wire#powerrail
      Contact( "T-103_SEQ_DB".RT_DATA.MOP.INIT )
      wire#w4
      I_Contact( "T-103_DB".Status.Aborting )
      Coil( "T-103_DB".Cmds.Abort )
   END_RUNG
   RUNG wire#powerrail
      Contact( "T-103_DB".Cmds.Abort )
   END_RUNG wire#w4
   // the same network as SCL:
   #_w1 := "T-103_HMI_DB".FromHMI.Stop OR "T-103_Read_FROM_R-201_DB".Aborting;
   #_w2 := #_w1 AND NOT "T-103_DB".OS.bit[0];   // rising edge
   "T-103_DB".OS.bit[0] := #_w1;
   "T-103_SEQ_DB".RT_DATA.MOP.INIT := #_w2 AND ((("T-103_SEQ_DB".S_NO > 1) AND NOT "T-103_DB".Status.Aborting) OR ("T-103_SEQ_DB".S_NO = 0));
   IF #_w2 THEN "T-103_HMI_DB".FromHMI.Stop := FALSE; END_IF;
   "T-103_DB".Cmds.Abort := ("T-103_SEQ_DB".RT_DATA.MOP.INIT OR "T-103_DB".Cmds.Abort) AND NOT "T-103_DB".Status.Aborting;
END_REGION

REGION Network 3: Initialize
   RUNG wire#powerrail
      Contact( "T-103_HMI_DB".FromHMI.Initialize )
      wire#w1
      I_Contact( "T-103_DB".Status.Aborting )
      I_Contact( "T-103_DB".Status.Running )
      wire#w2
      I_Contact( "T-103_DB".Status.Initializing )
      I_Contact( "T-103_DB".Cmds.Abort )
      I_Contact( "T-103_DB".Status.Ready )
      Coil( "T-103_DB".Cmds.Initialize )
   END_RUNG
   RUNG wire#powerrail
      Contact( "T-103_DB".ExchangeCmds.Receive.StartReceiving )
   END_RUNG wire#w1
   RUNG wire#powerrail
      Contact( "T-103_HMI_DB".FromHMI.Start )
      I_Contact( "T-103_DB".Cmds.Receive )
   END_RUNG wire#w1
   RUNG wire#powerrail
      Contact( "T-103_DB".Cmds.Initialize )
   END_RUNG wire#w2
   RUNG wire#powerrail
      Contact( "T-103_HMI_DB".FromHMI.Initialize )
      R_Coil( "T-103_HMI_DB".FromHMI.Initialize )
   END_RUNG
   // the same network as SCL:
   "T-103_DB".Cmds.Initialize := ((("T-103_HMI_DB".FromHMI.Initialize OR "T-103_DB".ExchangeCmds.Receive.StartReceiving OR ("T-103_HMI_DB".FromHMI.Start AND NOT "T-103_DB".Cmds.Receive)) AND NOT "T-103_DB".Status.Aborting AND NOT "T-103_DB".Status.Running) OR "T-103_DB".Cmds.Initialize) AND NOT "T-103_DB".Status.Initializing AND NOT "T-103_DB".Cmds.Abort AND NOT "T-103_DB".Status.Ready;
   IF "T-103_HMI_DB".FromHMI.Initialize THEN "T-103_HMI_DB".FromHMI.Initialize := FALSE; END_IF;
END_REGION

REGION Network 4: Start Receiving
   RUNG wire#powerrail
      Contact( "T-103_HMI_DB".FromHMI.Start )
      I_Contact( "T-103_DB".Status.Aborting )
      I_Contact( "T-103_DB".Status.Initializing )
      wire#w1
      I_Contact( "T-103_DB".Status.Running )
      I_Contact( "T-103_DB".Cmds.Abort )
      I_Contact( "T-103_DB".ExchangeCmds.Receive.StartReceiving )
      I_Contact( "T-103_DB".Cmds.Receive )
      Coil( "T-103_DB".Cmds.Start )
   END_RUNG
   RUNG wire#powerrail
      Contact( "T-103_DB".Cmds.Start )
   END_RUNG wire#w1
   RUNG wire#powerrail
      Contact( "T-103_HMI_DB".FromHMI.Start )
      R_Coil( "T-103_HMI_DB".FromHMI.Start )
   END_RUNG
   // the same network as SCL:
   "T-103_DB".Cmds.Start := (("T-103_HMI_DB".FromHMI.Start AND NOT "T-103_DB".Status.Aborting AND NOT "T-103_DB".Status.Initializing) OR "T-103_DB".Cmds.Start) AND NOT "T-103_DB".Status.Running AND NOT "T-103_DB".Cmds.Abort AND NOT "T-103_DB".ExchangeCmds.Receive.StartReceiving AND NOT "T-103_DB".Cmds.Receive;
   IF "T-103_HMI_DB".FromHMI.Start THEN "T-103_HMI_DB".FromHMI.Start := FALSE; END_IF;
END_REGION

